REGION Network 61
   RUNG wire#powerrail
      Move(in := "Carrier_03_CarrierDriveAlarm", out1 => "DB_SDC_EMS_TA".EMS[03].TA[1].ALARM)
      wire#w1
      Move(in := "Carrier_03_CarrierDriveAlarm", out1 => "EMS".Carrier[03].SDC_IN.CarrierDriveAlarms)
   END_RUNG
   RUNG wire#powerrail
      Contact( "IndiconTempDebugON" )
   END_RUNG wire#w1
   // the same network as SCL:
   "DB_SDC_EMS_TA".EMS[03].TA[1].ALARM := "Carrier_03_CarrierDriveAlarm";
   IF TRUE OR "IndiconTempDebugON" THEN
       "EMS".Carrier[03].SDC_IN.CarrierDriveAlarms := "Carrier_03_CarrierDriveAlarm";
   END_IF;
END_REGION

REGION Network 62
   RUNG wire#powerrail
      Move(in := "Carrier_03_SDCFaultCode", out1 => "DB101_DB_SDC_FAULTS".Carrier_Fault[03])
      wire#w1
      Move(in := "Carrier_03_SDCFaultCode", out1 => "EMS".Carrier[03].SDC_IN.CarrierFaults)
   END_RUNG
   RUNG wire#powerrail
      Contact( "IndiconTempDebugON" )
   END_RUNG wire#w1
   // the same network as SCL:
   "DB101_DB_SDC_FAULTS".Carrier_Fault[03] := "Carrier_03_SDCFaultCode";
   IF TRUE OR "IndiconTempDebugON" THEN
       "EMS".Carrier[03].SDC_IN.CarrierFaults := "Carrier_03_SDCFaultCode";
   END_IF;
END_REGION

REGION Network 63
   RUNG wire#powerrail
      Contact( "Carrier_03_Status.5" )
      Coil( "EMS".Carrier[03].SDC_IN.RunningFWD )
   END_RUNG
   // the same network as SCL:
   "EMS".Carrier[03].SDC_IN.RunningFWD := "Carrier_03_Status.5";
END_REGION

REGION Network 64
   RUNG wire#powerrail
      Contact( "Carrier_03_Status.6" )
      Coil( "EMS".Carrier[03].SDC_IN.RunningREV )
   END_RUNG
   // the same network as SCL:
   "EMS".Carrier[03].SDC_IN.RunningREV := "Carrier_03_Status.6";
END_REGION

REGION Network 65
   RUNG wire#powerrail
      Contact( "Carrier_03_Status.7" )
      Coil( "EMS".Carrier[03].SDC_IN.IR_Remote_9_Pressed )
   END_RUNG
   // the same network as SCL:
   "EMS".Carrier[03].SDC_IN.IR_Remote_9_Pressed := "Carrier_03_Status.7";
END_REGION

REGION Network 66
   RUNG wire#powerrail
      I_Contact( "Carrier_03_Status.5" )
      I_Contact( "Carrier_03_Status.6" )
      Coil( "EMS".Carrier[03].SDC_IN.Stopped )
   END_RUNG
   // the same network as SCL:
   "EMS".Carrier[03].SDC_IN.Stopped := NOT "Carrier_03_Status.5" AND NOT "Carrier_03_Status.6";
END_REGION

REGION Network 67
   RUNG wire#powerrail
      Contact( "Carrier_03_Status.4" )
      Coil( "EMS".Carrier[03].SDC_IN.ProductionHoldPB_Status )
   END_RUNG
   // the same network as SCL:
   "EMS".Carrier[03].SDC_IN.ProductionHoldPB_Status := "Carrier_03_Status.4";
END_REGION

REGION Network 68
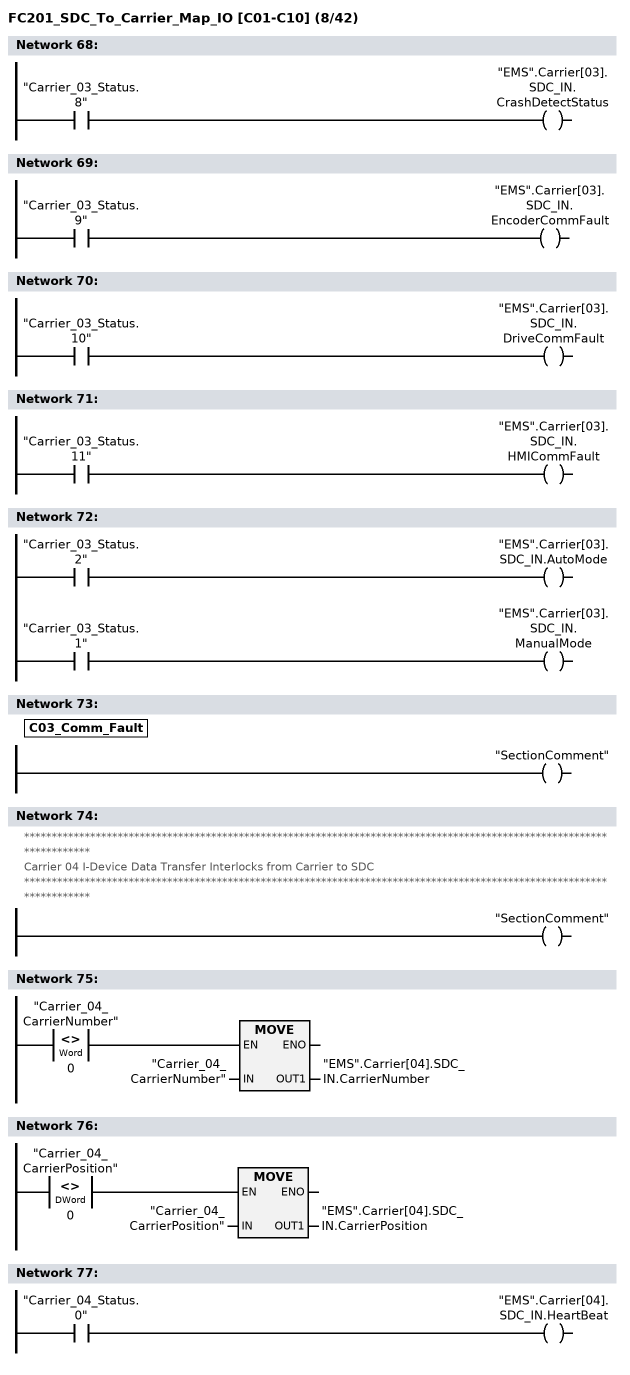
   RUNG wire#powerrail
      Contact( "Carrier_03_Status.8" )
      Coil( "EMS".Carrier[03].SDC_IN.CrashDetectStatus )
   END_RUNG
   // the same network as SCL:
   "EMS".Carrier[03].SDC_IN.CrashDetectStatus := "Carrier_03_Status.8";
END_REGION

REGION Network 69
   RUNG wire#powerrail
      Contact( "Carrier_03_Status.9" )
      Coil( "EMS".Carrier[03].SDC_IN.EncoderCommFault )
   END_RUNG
   // the same network as SCL:
   "EMS".Carrier[03].SDC_IN.EncoderCommFault := "Carrier_03_Status.9";
END_REGION

REGION Network 70
   RUNG wire#powerrail
      Contact( "Carrier_03_Status.10" )
      Coil( "EMS".Carrier[03].SDC_IN.DriveCommFault )
   END_RUNG
   // the same network as SCL:
   "EMS".Carrier[03].SDC_IN.DriveCommFault := "Carrier_03_Status.10";
END_REGION

REGION Network 71
   RUNG wire#powerrail
      Contact( "Carrier_03_Status.11" )
      Coil( "EMS".Carrier[03].SDC_IN.HMICommFault )
   END_RUNG
   // the same network as SCL:
   "EMS".Carrier[03].SDC_IN.HMICommFault := "Carrier_03_Status.11";
END_REGION

REGION Network 72
   RUNG wire#powerrail
      Contact( "Carrier_03_Status.2" )
      Coil( "EMS".Carrier[03].SDC_IN.AutoMode )
   END_RUNG
   RUNG wire#powerrail
      Contact( "Carrier_03_Status.1" )
      Coil( "EMS".Carrier[03].SDC_IN.ManualMode )
   END_RUNG
   // the same network as SCL:
   "EMS".Carrier[03].SDC_IN.AutoMode := "Carrier_03_Status.2";
   "EMS".Carrier[03].SDC_IN.ManualMode := "Carrier_03_Status.1";
END_REGION

REGION Network 73
   Label( C03_Comm_Fault )
   RUNG wire#powerrail
      Coil( "SectionComment" )
   END_RUNG
   // the same network as SCL:
   C03_Comm_Fault:
   "SectionComment" := TRUE;
END_REGION

REGION Network 74
   // **********************************************************************************************************************
   // 
   // Carrier 04 I-Device Data Transfer Interlocks from Carrier to SDC
   // 
   // **********************************************************************************************************************
   RUNG wire#powerrail
      Coil( "SectionComment" )
   END_RUNG
   // the same network as SCL:
   "SectionComment" := TRUE;
END_REGION

REGION Network 75
   RUNG wire#powerrail
      { S7_Templates := "SrcType := Word" } NE_Contact(in1 := "Carrier_04_CarrierNumber", in2 := 0)
      Move(in := "Carrier_04_CarrierNumber", out1 => "EMS".Carrier[04].SDC_IN.CarrierNumber)
   END_RUNG
   // the same network as SCL:
   IF "Carrier_04_CarrierNumber" <> 0 THEN
       "EMS".Carrier[04].SDC_IN.CarrierNumber := "Carrier_04_CarrierNumber";
   END_IF;
END_REGION

REGION Network 76
   RUNG wire#powerrail
      { S7_Templates := "SrcType := DWord" } NE_Contact(in1 := "Carrier_04_CarrierPosition", in2 := 0)
      Move(in := "Carrier_04_CarrierPosition", out1 => "EMS".Carrier[04].SDC_IN.CarrierPosition)
   END_RUNG
   // the same network as SCL:
   IF "Carrier_04_CarrierPosition" <> 0 THEN
       "EMS".Carrier[04].SDC_IN.CarrierPosition := "Carrier_04_CarrierPosition";
   END_IF;
END_REGION

REGION Network 77
   RUNG wire#powerrail
      Contact( "Carrier_04_Status.0" )
      Coil( "EMS".Carrier[04].SDC_IN.HeartBeat )
   END_RUNG
   // the same network as SCL:
   "EMS".Carrier[04].SDC_IN.HeartBeat := "Carrier_04_Status.0";
END_REGION

REGION Network 78
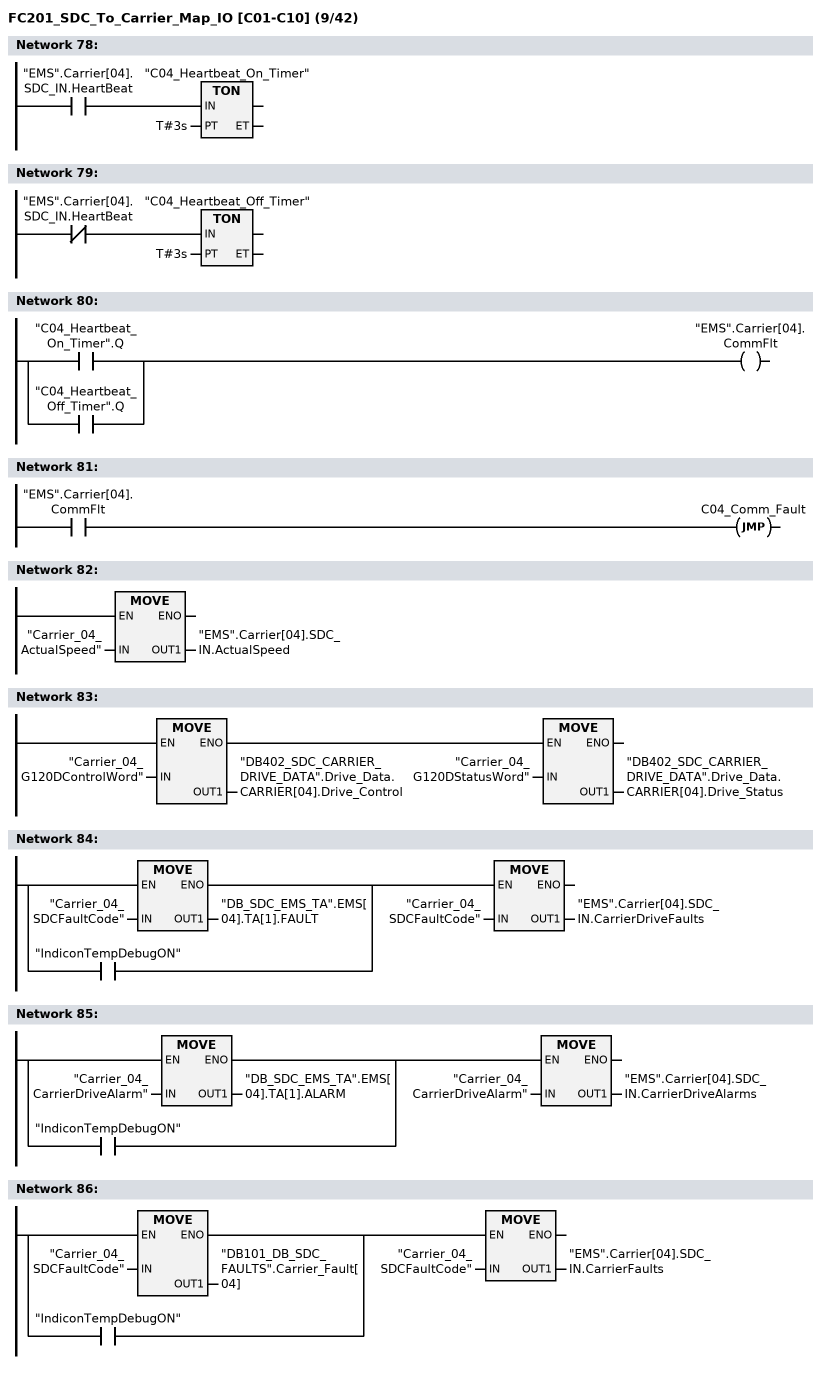
   "C04_Heartbeat_On_Timer".TON(IN := "EMS".Carrier[04].SDC_IN.HeartBeat, PT := T#3s);
END_REGION

REGION Network 79
   "C04_Heartbeat_Off_Timer".TON(IN := NOT "EMS".Carrier[04].SDC_IN.HeartBeat, PT := T#3s);
END_REGION

REGION Network 80
   RUNG wire#powerrail
      Contact( "C04_Heartbeat_On_Timer".Q )
      wire#w1
      Coil( "EMS".Carrier[04].CommFlt )
   END_RUNG
   RUNG wire#powerrail
      Contact( "C04_Heartbeat_Off_Timer".Q )
   END_RUNG wire#w1
   // the same network as SCL:
   "EMS".Carrier[04].CommFlt := "C04_Heartbeat_On_Timer".Q OR "C04_Heartbeat_Off_Timer".Q;
END_REGION

REGION Network 81
   RUNG wire#powerrail
      Contact( "EMS".Carrier[04].CommFlt )
      JumpCoil( C04_Comm_Fault )
   END_RUNG
   // the same network as SCL:
   IF "EMS".Carrier[04].CommFlt THEN GOTO C04_Comm_Fault; END_IF;
END_REGION

REGION Network 82
   RUNG wire#powerrail
      Move(in := "Carrier_04_ActualSpeed", out1 => "EMS".Carrier[04].SDC_IN.ActualSpeed)
   END_RUNG
   // the same network as SCL:
   "EMS".Carrier[04].SDC_IN.ActualSpeed := "Carrier_04_ActualSpeed";
END_REGION

REGION Network 83
   RUNG wire#powerrail
      Move(in := "Carrier_04_G120DControlWord", out1 => "DB402_SDC_CARRIER_DRIVE_DATA".Drive_Data.CARRIER[04].Drive_Control)
      Move(in := "Carrier_04_G120DStatusWord", out1 => "DB402_SDC_CARRIER_DRIVE_DATA".Drive_Data.CARRIER[04].Drive_Status)
   END_RUNG
   // the same network as SCL:
   "DB402_SDC_CARRIER_DRIVE_DATA".Drive_Data.CARRIER[04].Drive_Control := "Carrier_04_G120DControlWord";
   "DB402_SDC_CARRIER_DRIVE_DATA".Drive_Data.CARRIER[04].Drive_Status := "Carrier_04_G120DStatusWord";
END_REGION

REGION Network 84
   RUNG wire#powerrail
      Move(in := "Carrier_04_SDCFaultCode", out1 => "DB_SDC_EMS_TA".EMS[04].TA[1].FAULT)
      wire#w1
      Move(in := "Carrier_04_SDCFaultCode", out1 => "EMS".Carrier[04].SDC_IN.CarrierDriveFaults)
   END_RUNG
   RUNG wire#powerrail
      Contact( "IndiconTempDebugON" )
   END_RUNG wire#w1
   // the same network as SCL:
   "DB_SDC_EMS_TA".EMS[04].TA[1].FAULT := "Carrier_04_SDCFaultCode";
   IF TRUE OR "IndiconTempDebugON" THEN
       "EMS".Carrier[04].SDC_IN.CarrierDriveFaults := "Carrier_04_SDCFaultCode";
   END_IF;
END_REGION

REGION Network 85
   RUNG wire#powerrail
      Move(in := "Carrier_04_CarrierDriveAlarm", out1 => "DB_SDC_EMS_TA".EMS[04].TA[1].ALARM)
      wire#w1
      Move(in := "Carrier_04_CarrierDriveAlarm", out1 => "EMS".Carrier[04].SDC_IN.CarrierDriveAlarms)
   END_RUNG
   RUNG wire#powerrail
      Contact( "IndiconTempDebugON" )
   END_RUNG wire#w1
   // the same network as SCL:
   "DB_SDC_EMS_TA".EMS[04].TA[1].ALARM := "Carrier_04_CarrierDriveAlarm";
   IF TRUE OR "IndiconTempDebugON" THEN
       "EMS".Carrier[04].SDC_IN.CarrierDriveAlarms := "Carrier_04_CarrierDriveAlarm";
   END_IF;
END_REGION

REGION Network 86
   RUNG wire#powerrail
      Move(in := "Carrier_04_SDCFaultCode", out1 => "DB101_DB_SDC_FAULTS".Carrier_Fault[04])
      wire#w1
      Move(in := "Carrier_04_SDCFaultCode", out1 => "EMS".Carrier[04].SDC_IN.CarrierFaults)
   END_RUNG
   RUNG wire#powerrail
      Contact( "IndiconTempDebugON" )
   END_RUNG wire#w1
   // the same network as SCL:
   "DB101_DB_SDC_FAULTS".Carrier_Fault[04] := "Carrier_04_SDCFaultCode";
   IF TRUE OR "IndiconTempDebugON" THEN
       "EMS".Carrier[04].SDC_IN.CarrierFaults := "Carrier_04_SDCFaultCode";
   END_IF;
END_REGION

REGION Network 87
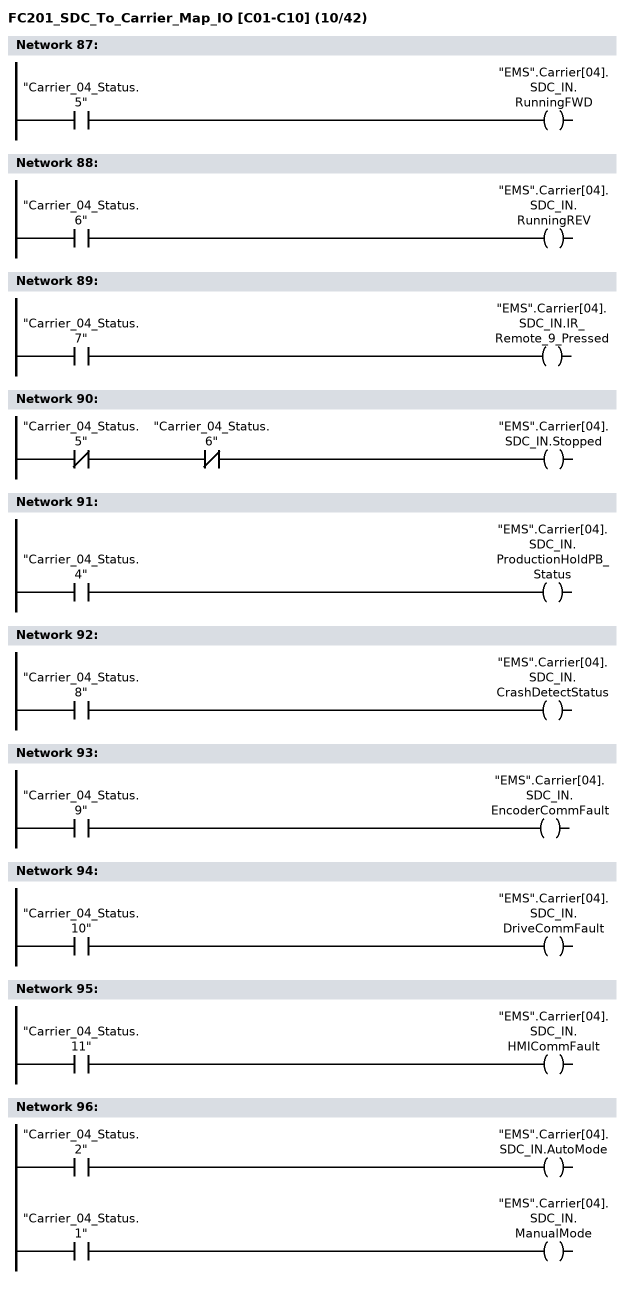
   RUNG wire#powerrail
      Contact( "Carrier_04_Status.5" )
      Coil( "EMS".Carrier[04].SDC_IN.RunningFWD )
   END_RUNG
   // the same network as SCL:
   "EMS".Carrier[04].SDC_IN.RunningFWD := "Carrier_04_Status.5";
END_REGION

REGION Network 88
   RUNG wire#powerrail
      Contact( "Carrier_04_Status.6" )
      Coil( "EMS".Carrier[04].SDC_IN.RunningREV )
   END_RUNG
   // the same network as SCL:
   "EMS".Carrier[04].SDC_IN.RunningREV := "Carrier_04_Status.6";
END_REGION

REGION Network 89
   RUNG wire#powerrail
      Contact( "Carrier_04_Status.7" )
      Coil( "EMS".Carrier[04].SDC_IN.IR_Remote_9_Pressed )
   END_RUNG
   // the same network as SCL:
   "EMS".Carrier[04].SDC_IN.IR_Remote_9_Pressed := "Carrier_04_Status.7";
END_REGION

REGION Network 90
   RUNG wire#powerrail
      I_Contact( "Carrier_04_Status.5" )
      I_Contact( "Carrier_04_Status.6" )
      Coil( "EMS".Carrier[04].SDC_IN.Stopped )
   END_RUNG
   // the same network as SCL:
   "EMS".Carrier[04].SDC_IN.Stopped := NOT "Carrier_04_Status.5" AND NOT "Carrier_04_Status.6";
END_REGION

REGION Network 91
   RUNG wire#powerrail
      Contact( "Carrier_04_Status.4" )
      Coil( "EMS".Carrier[04].SDC_IN.ProductionHoldPB_Status )
   END_RUNG
   // the same network as SCL:
   "EMS".Carrier[04].SDC_IN.ProductionHoldPB_Status := "Carrier_04_Status.4";
END_REGION

REGION Network 92
   RUNG wire#powerrail
      Contact( "Carrier_04_Status.8" )
      Coil( "EMS".Carrier[04].SDC_IN.CrashDetectStatus )
   END_RUNG
   // the same network as SCL:
   "EMS".Carrier[04].SDC_IN.CrashDetectStatus := "Carrier_04_Status.8";
END_REGION

REGION Network 93
   RUNG wire#powerrail
      Contact( "Carrier_04_Status.9" )
      Coil( "EMS".Carrier[04].SDC_IN.EncoderCommFault )
   END_RUNG
   // the same network as SCL:
   "EMS".Carrier[04].SDC_IN.EncoderCommFault := "Carrier_04_Status.9";
END_REGION

REGION Network 94
   RUNG wire#powerrail
      Contact( "Carrier_04_Status.10" )
      Coil( "EMS".Carrier[04].SDC_IN.DriveCommFault )
   END_RUNG
   // the same network as SCL:
   "EMS".Carrier[04].SDC_IN.DriveCommFault := "Carrier_04_Status.10";
END_REGION

REGION Network 95
   RUNG wire#powerrail
      Contact( "Carrier_04_Status.11" )
      Coil( "EMS".Carrier[04].SDC_IN.HMICommFault )
   END_RUNG
   // the same network as SCL:
   "EMS".Carrier[04].SDC_IN.HMICommFault := "Carrier_04_Status.11";
END_REGION

REGION Network 96
   RUNG wire#powerrail
      Contact( "Carrier_04_Status.2" )
      Coil( "EMS".Carrier[04].SDC_IN.AutoMode )
   END_RUNG
   RUNG wire#powerrail
      Contact( "Carrier_04_Status.1" )
      Coil( "EMS".Carrier[04].SDC_IN.ManualMode )
   END_RUNG
   // the same network as SCL:
   "EMS".Carrier[04].SDC_IN.AutoMode := "Carrier_04_Status.2";
   "EMS".Carrier[04].SDC_IN.ManualMode := "Carrier_04_Status.1";
END_REGION

REGION Network 97
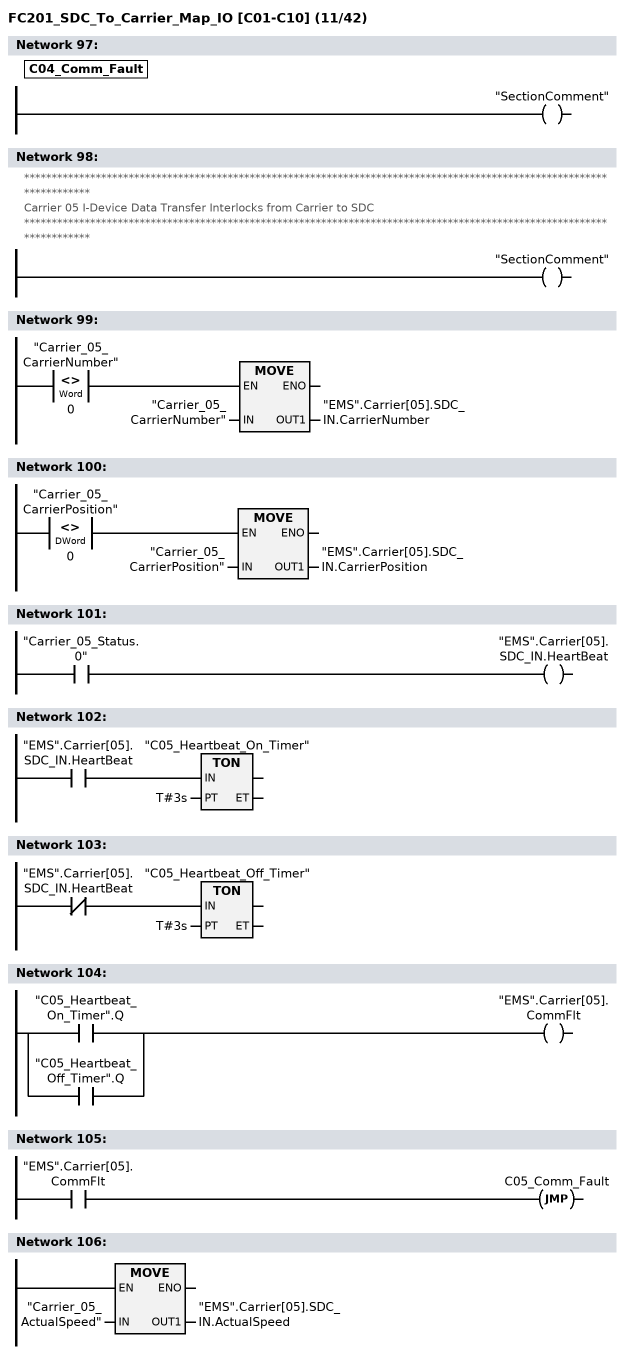
   Label( C04_Comm_Fault )
   RUNG wire#powerrail
      Coil( "SectionComment" )
   END_RUNG
   // the same network as SCL:
   C04_Comm_Fault:
   "SectionComment" := TRUE;
END_REGION

REGION Network 98
   // **********************************************************************************************************************
   // 
   // Carrier 05 I-Device Data Transfer Interlocks from Carrier to SDC
   // 
   // **********************************************************************************************************************
   RUNG wire#powerrail
      Coil( "SectionComment" )
   END_RUNG
   // the same network as SCL:
   "SectionComment" := TRUE;
END_REGION

REGION Network 99
   RUNG wire#powerrail
      { S7_Templates := "SrcType := Word" } NE_Contact(in1 := "Carrier_05_CarrierNumber", in2 := 0)
      Move(in := "Carrier_05_CarrierNumber", out1 => "EMS".Carrier[05].SDC_IN.CarrierNumber)
   END_RUNG
   // the same network as SCL:
   IF "Carrier_05_CarrierNumber" <> 0 THEN
       "EMS".Carrier[05].SDC_IN.CarrierNumber := "Carrier_05_CarrierNumber";
   END_IF;
END_REGION

REGION Network 100
   RUNG wire#powerrail
      { S7_Templates := "SrcType := DWord" } NE_Contact(in1 := "Carrier_05_CarrierPosition", in2 := 0)
      Move(in := "Carrier_05_CarrierPosition", out1 => "EMS".Carrier[05].SDC_IN.CarrierPosition)
   END_RUNG
   // the same network as SCL:
   IF "Carrier_05_CarrierPosition" <> 0 THEN
       "EMS".Carrier[05].SDC_IN.CarrierPosition := "Carrier_05_CarrierPosition";
   END_IF;
END_REGION

REGION Network 101
   RUNG wire#powerrail
      Contact( "Carrier_05_Status.0" )
      Coil( "EMS".Carrier[05].SDC_IN.HeartBeat )
   END_RUNG
   // the same network as SCL:
   "EMS".Carrier[05].SDC_IN.HeartBeat := "Carrier_05_Status.0";
END_REGION

REGION Network 102
   "C05_Heartbeat_On_Timer".TON(IN := "EMS".Carrier[05].SDC_IN.HeartBeat, PT := T#3s);
END_REGION

REGION Network 103
   "C05_Heartbeat_Off_Timer".TON(IN := NOT "EMS".Carrier[05].SDC_IN.HeartBeat, PT := T#3s);
END_REGION

REGION Network 104
   RUNG wire#powerrail
      Contact( "C05_Heartbeat_On_Timer".Q )
      wire#w1
      Coil( "EMS".Carrier[05].CommFlt )
   END_RUNG
   RUNG wire#powerrail
      Contact( "C05_Heartbeat_Off_Timer".Q )
   END_RUNG wire#w1
   // the same network as SCL:
   "EMS".Carrier[05].CommFlt := "C05_Heartbeat_On_Timer".Q OR "C05_Heartbeat_Off_Timer".Q;
END_REGION

REGION Network 105
   RUNG wire#powerrail
      Contact( "EMS".Carrier[05].CommFlt )
      JumpCoil( C05_Comm_Fault )
   END_RUNG
   // the same network as SCL:
   IF "EMS".Carrier[05].CommFlt THEN GOTO C05_Comm_Fault; END_IF;
END_REGION

REGION Network 106
   RUNG wire#powerrail
      Move(in := "Carrier_05_ActualSpeed", out1 => "EMS".Carrier[05].SDC_IN.ActualSpeed)
   END_RUNG
   // the same network as SCL:
   "EMS".Carrier[05].SDC_IN.ActualSpeed := "Carrier_05_ActualSpeed";
END_REGION

REGION Network 107
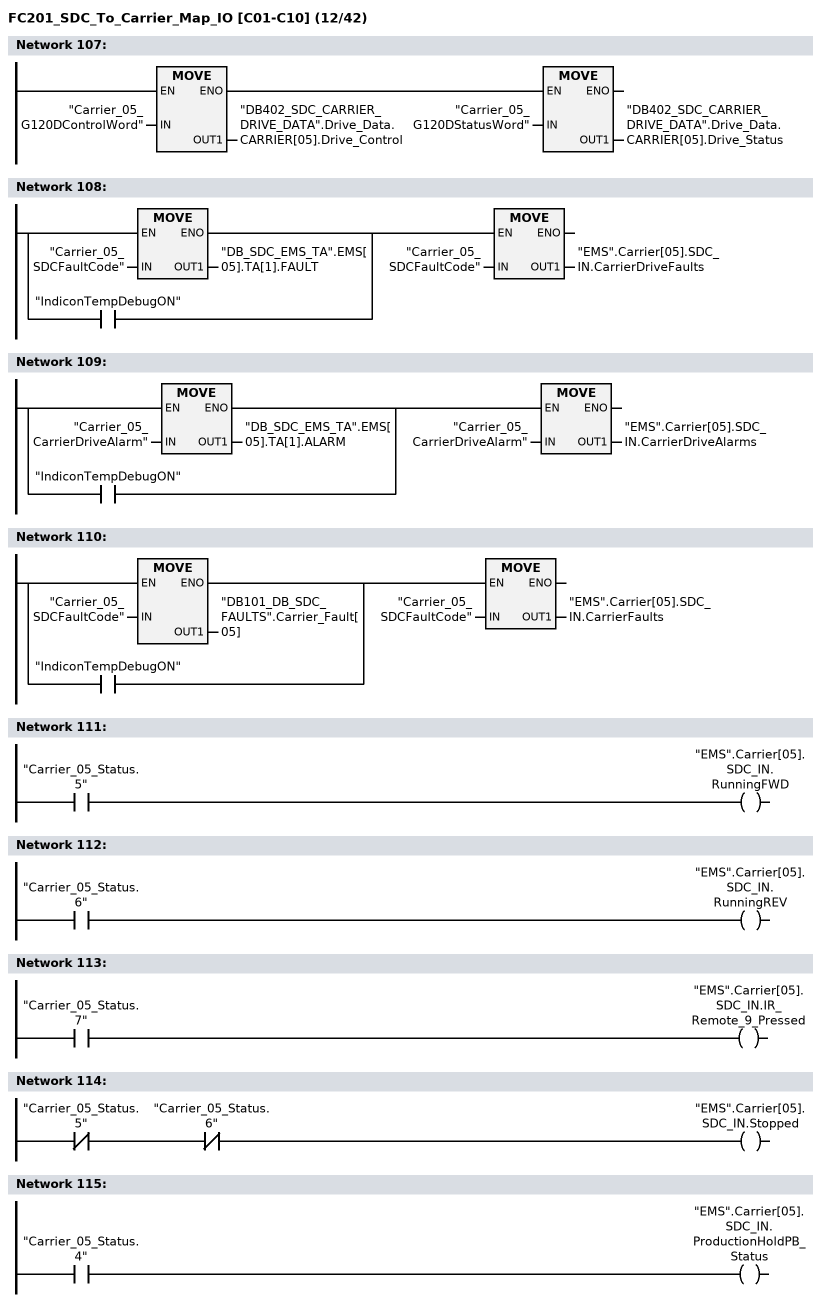
   RUNG wire#powerrail
      Move(in := "Carrier_05_G120DControlWord", out1 => "DB402_SDC_CARRIER_DRIVE_DATA".Drive_Data.CARRIER[05].Drive_Control)
      Move(in := "Carrier_05_G120DStatusWord", out1 => "DB402_SDC_CARRIER_DRIVE_DATA".Drive_Data.CARRIER[05].Drive_Status)
   END_RUNG
   // the same network as SCL:
   "DB402_SDC_CARRIER_DRIVE_DATA".Drive_Data.CARRIER[05].Drive_Control := "Carrier_05_G120DControlWord";
   "DB402_SDC_CARRIER_DRIVE_DATA".Drive_Data.CARRIER[05].Drive_Status := "Carrier_05_G120DStatusWord";
END_REGION

REGION Network 108
   RUNG wire#powerrail
      Move(in := "Carrier_05_SDCFaultCode", out1 => "DB_SDC_EMS_TA".EMS[05].TA[1].FAULT)
      wire#w1
      Move(in := "Carrier_05_SDCFaultCode", out1 => "EMS".Carrier[05].SDC_IN.CarrierDriveFaults)
   END_RUNG
   RUNG wire#powerrail
      Contact( "IndiconTempDebugON" )
   END_RUNG wire#w1
   // the same network as SCL:
   "DB_SDC_EMS_TA".EMS[05].TA[1].FAULT := "Carrier_05_SDCFaultCode";
   IF TRUE OR "IndiconTempDebugON" THEN
       "EMS".Carrier[05].SDC_IN.CarrierDriveFaults := "Carrier_05_SDCFaultCode";
   END_IF;
END_REGION

REGION Network 109
   RUNG wire#powerrail
      Move(in := "Carrier_05_CarrierDriveAlarm", out1 => "DB_SDC_EMS_TA".EMS[05].TA[1].ALARM)
      wire#w1
      Move(in := "Carrier_05_CarrierDriveAlarm", out1 => "EMS".Carrier[05].SDC_IN.CarrierDriveAlarms)
   END_RUNG
   RUNG wire#powerrail
      Contact( "IndiconTempDebugON" )
   END_RUNG wire#w1
   // the same network as SCL:
   "DB_SDC_EMS_TA".EMS[05].TA[1].ALARM := "Carrier_05_CarrierDriveAlarm";
   IF TRUE OR "IndiconTempDebugON" THEN
       "EMS".Carrier[05].SDC_IN.CarrierDriveAlarms := "Carrier_05_CarrierDriveAlarm";
   END_IF;
END_REGION

REGION Network 110
   RUNG wire#powerrail
      Move(in := "Carrier_05_SDCFaultCode", out1 => "DB101_DB_SDC_FAULTS".Carrier_Fault[05])
      wire#w1
      Move(in := "Carrier_05_SDCFaultCode", out1 => "EMS".Carrier[05].SDC_IN.CarrierFaults)
   END_RUNG
   RUNG wire#powerrail
      Contact( "IndiconTempDebugON" )
   END_RUNG wire#w1
   // the same network as SCL:
   "DB101_DB_SDC_FAULTS".Carrier_Fault[05] := "Carrier_05_SDCFaultCode";
   IF TRUE OR "IndiconTempDebugON" THEN
       "EMS".Carrier[05].SDC_IN.CarrierFaults := "Carrier_05_SDCFaultCode";
   END_IF;
END_REGION

REGION Network 111
   RUNG wire#powerrail
      Contact( "Carrier_05_Status.5" )
      Coil( "EMS".Carrier[05].SDC_IN.RunningFWD )
   END_RUNG
   // the same network as SCL:
   "EMS".Carrier[05].SDC_IN.RunningFWD := "Carrier_05_Status.5";
END_REGION

REGION Network 112
   RUNG wire#powerrail
      Contact( "Carrier_05_Status.6" )
      Coil( "EMS".Carrier[05].SDC_IN.RunningREV )
   END_RUNG
   // the same network as SCL:
   "EMS".Carrier[05].SDC_IN.RunningREV := "Carrier_05_Status.6";
END_REGION

REGION Network 113
   RUNG wire#powerrail
      Contact( "Carrier_05_Status.7" )
      Coil( "EMS".Carrier[05].SDC_IN.IR_Remote_9_Pressed )
   END_RUNG
   // the same network as SCL:
   "EMS".Carrier[05].SDC_IN.IR_Remote_9_Pressed := "Carrier_05_Status.7";
END_REGION

REGION Network 114
   RUNG wire#powerrail
      I_Contact( "Carrier_05_Status.5" )
      I_Contact( "Carrier_05_Status.6" )
      Coil( "EMS".Carrier[05].SDC_IN.Stopped )
   END_RUNG
   // the same network as SCL:
   "EMS".Carrier[05].SDC_IN.Stopped := NOT "Carrier_05_Status.5" AND NOT "Carrier_05_Status.6";
END_REGION

REGION Network 115
   RUNG wire#powerrail
      Contact( "Carrier_05_Status.4" )
      Coil( "EMS".Carrier[05].SDC_IN.ProductionHoldPB_Status )
   END_RUNG
   // the same network as SCL:
   "EMS".Carrier[05].SDC_IN.ProductionHoldPB_Status := "Carrier_05_Status.4";
END_REGION

REGION Network 116
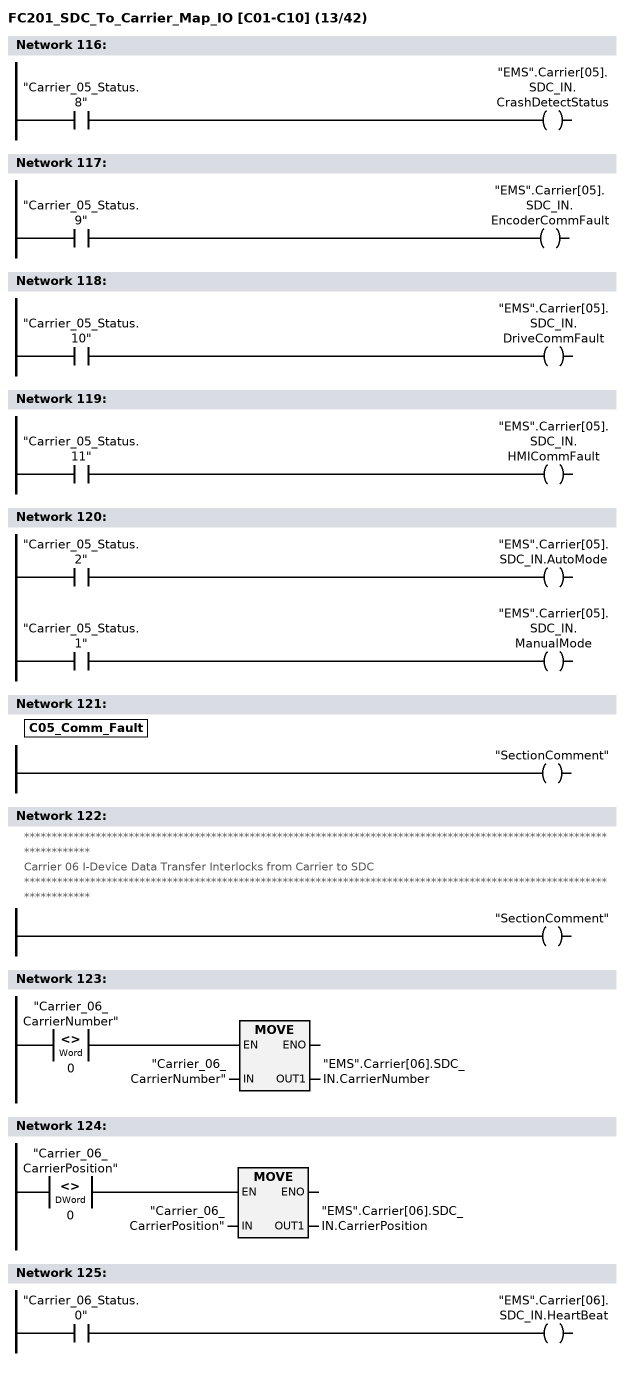
   RUNG wire#powerrail
      Contact( "Carrier_05_Status.8" )
      Coil( "EMS".Carrier[05].SDC_IN.CrashDetectStatus )
   END_RUNG
   // the same network as SCL:
   "EMS".Carrier[05].SDC_IN.CrashDetectStatus := "Carrier_05_Status.8";
END_REGION

REGION Network 117
   RUNG wire#powerrail
      Contact( "Carrier_05_Status.9" )
      Coil( "EMS".Carrier[05].SDC_IN.EncoderCommFault )
   END_RUNG
   // the same network as SCL:
   "EMS".Carrier[05].SDC_IN.EncoderCommFault := "Carrier_05_Status.9";
END_REGION

REGION Network 118
   RUNG wire#powerrail
      Contact( "Carrier_05_Status.10" )
      Coil( "EMS".Carrier[05].SDC_IN.DriveCommFault )
   END_RUNG
   // the same network as SCL:
   "EMS".Carrier[05].SDC_IN.DriveCommFault := "Carrier_05_Status.10";
END_REGION

REGION Network 119
   RUNG wire#powerrail
      Contact( "Carrier_05_Status.11" )
      Coil( "EMS".Carrier[05].SDC_IN.HMICommFault )
   END_RUNG
   // the same network as SCL:
   "EMS".Carrier[05].SDC_IN.HMICommFault := "Carrier_05_Status.11";
END_REGION

REGION Network 120
   RUNG wire#powerrail
      Contact( "Carrier_05_Status.2" )
      Coil( "EMS".Carrier[05].SDC_IN.AutoMode )
   END_RUNG
   RUNG wire#powerrail
      Contact( "Carrier_05_Status.1" )
      Coil( "EMS".Carrier[05].SDC_IN.ManualMode )
   END_RUNG
   // the same network as SCL:
   "EMS".Carrier[05].SDC_IN.AutoMode := "Carrier_05_Status.2";
   "EMS".Carrier[05].SDC_IN.ManualMode := "Carrier_05_Status.1";
END_REGION

REGION Network 121
   Label( C05_Comm_Fault )
   RUNG wire#powerrail
      Coil( "SectionComment" )
   END_RUNG
   // the same network as SCL:
   C05_Comm_Fault:
   "SectionComment" := TRUE;
END_REGION

REGION Network 122
   // **********************************************************************************************************************
   // 
   // Carrier 06 I-Device Data Transfer Interlocks from Carrier to SDC
   // 
   // **********************************************************************************************************************
   RUNG wire#powerrail
      Coil( "SectionComment" )
   END_RUNG
   // the same network as SCL:
   "SectionComment" := TRUE;
END_REGION

REGION Network 123
   RUNG wire#powerrail
      { S7_Templates := "SrcType := Word" } NE_Contact(in1 := "Carrier_06_CarrierNumber", in2 := 0)
      Move(in := "Carrier_06_CarrierNumber", out1 => "EMS".Carrier[06].SDC_IN.CarrierNumber)
   END_RUNG
   // the same network as SCL:
   IF "Carrier_06_CarrierNumber" <> 0 THEN
       "EMS".Carrier[06].SDC_IN.CarrierNumber := "Carrier_06_CarrierNumber";
   END_IF;
END_REGION

REGION Network 124
   RUNG wire#powerrail
      { S7_Templates := "SrcType := DWord" } NE_Contact(in1 := "Carrier_06_CarrierPosition", in2 := 0)
      Move(in := "Carrier_06_CarrierPosition", out1 => "EMS".Carrier[06].SDC_IN.CarrierPosition)
   END_RUNG
   // the same network as SCL:
   IF "Carrier_06_CarrierPosition" <> 0 THEN
       "EMS".Carrier[06].SDC_IN.CarrierPosition := "Carrier_06_CarrierPosition";
   END_IF;
END_REGION

REGION Network 125
   RUNG wire#powerrail
      Contact( "Carrier_06_Status.0" )
      Coil( "EMS".Carrier[06].SDC_IN.HeartBeat )
   END_RUNG
   // the same network as SCL:
   "EMS".Carrier[06].SDC_IN.HeartBeat := "Carrier_06_Status.0";
END_REGION

REGION Network 126
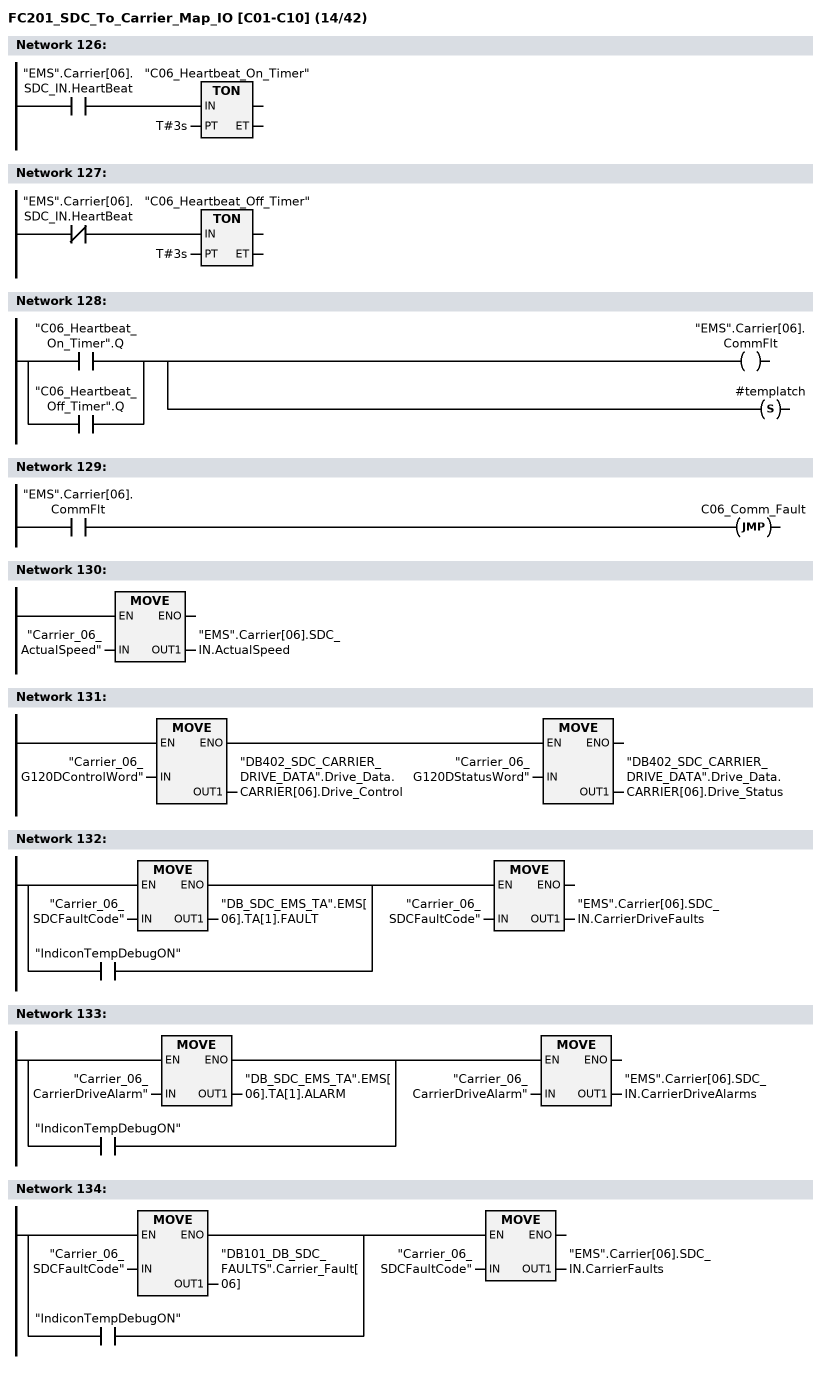
   "C06_Heartbeat_On_Timer".TON(IN := "EMS".Carrier[06].SDC_IN.HeartBeat, PT := T#3s);
END_REGION

REGION Network 127
   "C06_Heartbeat_Off_Timer".TON(IN := NOT "EMS".Carrier[06].SDC_IN.HeartBeat, PT := T#3s);
END_REGION

REGION Network 128
   RUNG wire#powerrail
      Contact( "C06_Heartbeat_On_Timer".Q )
      wire#w1
      Coil( "EMS".Carrier[06].CommFlt )
   END_RUNG
   RUNG wire#powerrail
      Contact( "C06_Heartbeat_Off_Timer".Q )
   END_RUNG wire#w1
   RUNG wire#w1
      S_Coil( #templatch )
   END_RUNG
   // the same network as SCL:
   "EMS".Carrier[06].CommFlt := "C06_Heartbeat_On_Timer".Q OR "C06_Heartbeat_Off_Timer".Q;
   IF "C06_Heartbeat_On_Timer".Q OR "C06_Heartbeat_Off_Timer".Q THEN #templatch := TRUE; END_IF;
END_REGION

REGION Network 129
   RUNG wire#powerrail
      Contact( "EMS".Carrier[06].CommFlt )
      JumpCoil( C06_Comm_Fault )
   END_RUNG
   // the same network as SCL:
   IF "EMS".Carrier[06].CommFlt THEN GOTO C06_Comm_Fault; END_IF;
END_REGION

REGION Network 130
   RUNG wire#powerrail
      Move(in := "Carrier_06_ActualSpeed", out1 => "EMS".Carrier[06].SDC_IN.ActualSpeed)
   END_RUNG
   // the same network as SCL:
   "EMS".Carrier[06].SDC_IN.ActualSpeed := "Carrier_06_ActualSpeed";
END_REGION

REGION Network 131
   RUNG wire#powerrail
      Move(in := "Carrier_06_G120DControlWord", out1 => "DB402_SDC_CARRIER_DRIVE_DATA".Drive_Data.CARRIER[06].Drive_Control)
      Move(in := "Carrier_06_G120DStatusWord", out1 => "DB402_SDC_CARRIER_DRIVE_DATA".Drive_Data.CARRIER[06].Drive_Status)
   END_RUNG
   // the same network as SCL:
   "DB402_SDC_CARRIER_DRIVE_DATA".Drive_Data.CARRIER[06].Drive_Control := "Carrier_06_G120DControlWord";
   "DB402_SDC_CARRIER_DRIVE_DATA".Drive_Data.CARRIER[06].Drive_Status := "Carrier_06_G120DStatusWord";
END_REGION

REGION Network 132
   RUNG wire#powerrail
      Move(in := "Carrier_06_SDCFaultCode", out1 => "DB_SDC_EMS_TA".EMS[06].TA[1].FAULT)
      wire#w1
      Move(in := "Carrier_06_SDCFaultCode", out1 => "EMS".Carrier[06].SDC_IN.CarrierDriveFaults)
   END_RUNG
   RUNG wire#powerrail
      Contact( "IndiconTempDebugON" )
   END_RUNG wire#w1
   // the same network as SCL:
   "DB_SDC_EMS_TA".EMS[06].TA[1].FAULT := "Carrier_06_SDCFaultCode";
   IF TRUE OR "IndiconTempDebugON" THEN
       "EMS".Carrier[06].SDC_IN.CarrierDriveFaults := "Carrier_06_SDCFaultCode";
   END_IF;
END_REGION

REGION Network 133
   RUNG wire#powerrail
      Move(in := "Carrier_06_CarrierDriveAlarm", out1 => "DB_SDC_EMS_TA".EMS[06].TA[1].ALARM)
      wire#w1
      Move(in := "Carrier_06_CarrierDriveAlarm", out1 => "EMS".Carrier[06].SDC_IN.CarrierDriveAlarms)
   END_RUNG
   RUNG wire#powerrail
      Contact( "IndiconTempDebugON" )
   END_RUNG wire#w1
   // the same network as SCL:
   "DB_SDC_EMS_TA".EMS[06].TA[1].ALARM := "Carrier_06_CarrierDriveAlarm";
   IF TRUE OR "IndiconTempDebugON" THEN
       "EMS".Carrier[06].SDC_IN.CarrierDriveAlarms := "Carrier_06_CarrierDriveAlarm";
   END_IF;
END_REGION

REGION Network 134
   RUNG wire#powerrail
      Move(in := "Carrier_06_SDCFaultCode", out1 => "DB101_DB_SDC_FAULTS".Carrier_Fault[06])
      wire#w1
      Move(in := "Carrier_06_SDCFaultCode", out1 => "EMS".Carrier[06].SDC_IN.CarrierFaults)
   END_RUNG
   RUNG wire#powerrail
      Contact( "IndiconTempDebugON" )
   END_RUNG wire#w1
   // the same network as SCL:
   "DB101_DB_SDC_FAULTS".Carrier_Fault[06] := "Carrier_06_SDCFaultCode";
   IF TRUE OR "IndiconTempDebugON" THEN
       "EMS".Carrier[06].SDC_IN.CarrierFaults := "Carrier_06_SDCFaultCode";
   END_IF;
END_REGION

REGION Network 135
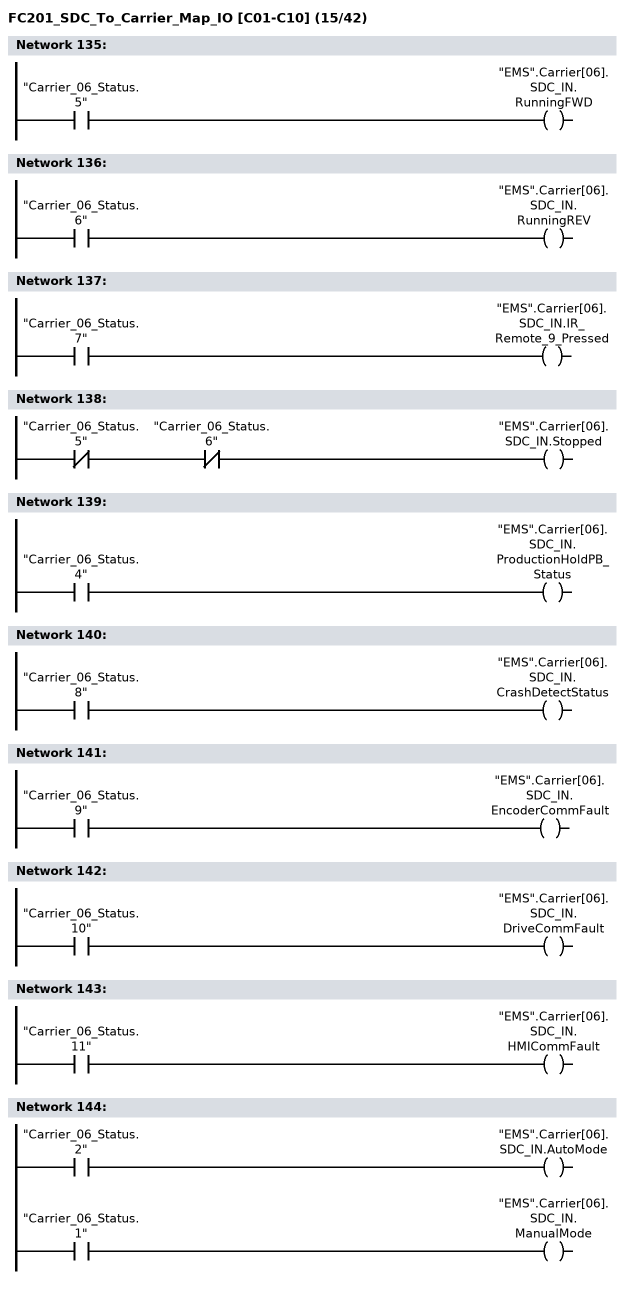
   RUNG wire#powerrail
      Contact( "Carrier_06_Status.5" )
      Coil( "EMS".Carrier[06].SDC_IN.RunningFWD )
   END_RUNG
   // the same network as SCL:
   "EMS".Carrier[06].SDC_IN.RunningFWD := "Carrier_06_Status.5";
END_REGION

REGION Network 136
   RUNG wire#powerrail
      Contact( "Carrier_06_Status.6" )
      Coil( "EMS".Carrier[06].SDC_IN.RunningREV )
   END_RUNG
   // the same network as SCL:
   "EMS".Carrier[06].SDC_IN.RunningREV := "Carrier_06_Status.6";
END_REGION

REGION Network 137
   RUNG wire#powerrail
      Contact( "Carrier_06_Status.7" )
      Coil( "EMS".Carrier[06].SDC_IN.IR_Remote_9_Pressed )
   END_RUNG
   // the same network as SCL:
   "EMS".Carrier[06].SDC_IN.IR_Remote_9_Pressed := "Carrier_06_Status.7";
END_REGION

REGION Network 138
   RUNG wire#powerrail
      I_Contact( "Carrier_06_Status.5" )
      I_Contact( "Carrier_06_Status.6" )
      Coil( "EMS".Carrier[06].SDC_IN.Stopped )
   END_RUNG
   // the same network as SCL:
   "EMS".Carrier[06].SDC_IN.Stopped := NOT "Carrier_06_Status.5" AND NOT "Carrier_06_Status.6";
END_REGION

REGION Network 139
   RUNG wire#powerrail
      Contact( "Carrier_06_Status.4" )
      Coil( "EMS".Carrier[06].SDC_IN.ProductionHoldPB_Status )
   END_RUNG
   // the same network as SCL:
   "EMS".Carrier[06].SDC_IN.ProductionHoldPB_Status := "Carrier_06_Status.4";
END_REGION

REGION Network 140
   RUNG wire#powerrail
      Contact( "Carrier_06_Status.8" )
      Coil( "EMS".Carrier[06].SDC_IN.CrashDetectStatus )
   END_RUNG
   // the same network as SCL:
   "EMS".Carrier[06].SDC_IN.CrashDetectStatus := "Carrier_06_Status.8";
END_REGION
